VERSION : 0.7
   VAR_INPUT
      FB_Mode : Int;   // Function Block Mode - 0 = HOA Directly Wired to SMC / 1 = HOA Remotely Wired
      MANM : Bool;   // Used only for FB_Mode = 1 / Manual Mode Signal
      AUTM : Bool;   // Used only for FB_Mode = 1 / Auto Mode Signal
      IL : Bool;   // Interlock
      HON : Bool;   // Hand ON
      HOFF : Bool;   // Hand OFF
      SpareIN_1 : Bool;   // Spare
      SRM : Bool;   // Status - Remote Mode Feedback
      SON : Bool;   // Status - On
      SDO : Bool;   // Status - Device Ok
      SCDPA : Bool;   // Status - Cooling Down Period Active
      SESE : Bool;   // Status - Emergency Start Executed
      SGW : Bool;   // Fault - General Warning
      SGF : Bool;   // Fault - General Fault
      EOLO : Bool;   // Event - Overload Operation Fault (I>115%Is)
      EOL : Bool;   // Event - Overload Fault
      EUN : Bool;   // Event - Unbalance Fault
      EOLLP : Bool;   // Event - Overload and Loss of Phase
      ESR : Bool;   // Event - Stalled Rotor
      THFBU : Bool;   // Trip - Hardware Fault Basic Unit
      TMF : Bool;   // Trip - Module Fault
      TEOC : Bool;   // Trip - Execution On-Command
      MC : Int;   // Maximum Current (% of Is)
      IL1 : Int;   // Current of Leg 1 (% of Is)
      IL2 : Int;   // Current of Leg 2 (% of Is)
      IL3 : Int;   // Current of Leg 3 (% of Is)
      RCDP : Int;   // Remaining Cool Down Period
      MOHH : Int;   // Motor Operating Hours High Word
      MOHL : Int;   // Motor Operating Hours Low Word
      LTC : Int;   // Last Trip Current (% of Is)
      "NOT" : Int;   // Number of Overload Trips
      FLA : Real;   // Full Load Amps
   END_VAR
   VAR_OUTPUT
      SpareOUT_1 : Bool;
      Stop_CMD : Bool;   // Stop Command for the Semicode
      Start_CMD : Bool;   // Start Command for the Semicode
      TST : Bool;   // Simocode Test
      EST : Bool;   // Emergency Start
      ERC : Bool;   // Auto Mode / Enable Remote Commands
      RST : Bool;   // Simocode Reset
      SpareOUT_2 : Bool;
      SpareOUT_3 : Bool;
      SpareOUT_4 : Bool;
      SpareOUT_5 : Bool;
      SpareOUT_6 : Bool;
      SpareOUT_7 : Bool;
      SpareOUT_8 : Bool;
      SpareOUT_9 : Bool;
      SpareOUT_10 : Bool;
      SpareOUTW_1 : Int;
      SpareOUTW_2 : Int;
   END_VAR
   VAR
      HMI : Struct
         Controls : Struct
            Start : Bool;
            Stop : Bool;
            Reset : Bool;
            PLCMOHR : Bool;   // PLC Motor Operating Hours Reset
         END_STRUCT;
         Status : Struct
            Mode : Int;   // Simocode Mode
            MotorOperatingHours : Real;   // True Semicode Motor Operating Hours
            DeviceOperatingHours : Real;
            LMOH : Real;   // Last Motor Operating Hours
            RemainingCoolDownPeriod : Int;   // Remaining Cooldown Period
            MaxNumberOLtrips : Int;   // Maximum Number of Overload Trips
            ControlStatusWord : Word;   // Control/Status Information Bits
            MaxCurrent : Real;   // Maximum Current (Is %)
            Current1 : Real;   // Leg 1 Current (Is %)
            Current2 : Real;   // Leg 2 Current (Is %)
            Current3 : Real;   // Leg 3 Current (Is %)
            LastTripCurrent : Real;   // Last Trip Current (% of Is)
            CommandSimocode : Bool;   // Commanding Simocode to Start
         END_STRUCT;
         Config : Struct
            "RemainingCoolDownPeriod.SP" : Int := 300;
            Start_PT : Time := T#500MS;
            Stop_PT : Time := T#500MS;
         END_STRUCT;
         Math : Struct
            MOH1 : DInt;
            MOH2 : Real;
            PLCMOH : Real;   // PLC Motor Operating Hours
            LMOH : Real;
         END_STRUCT;
      END_STRUCT;
      OS : Struct
         RON : Bool;   // Remote / HMI On
         ROFF : Bool;   // Remote / HMI Off
         HON : Bool;   // Hand/Local On
         HOFF : Bool;   // Hand/Local Off
         PLCMOHR : Bool;
         LMOH1 : Bool;
         LMOH2 : Bool;
         RST : Bool;   // Reset Semicode
      END_STRUCT;
      START_CMD_TOF : TOF_TIME;   // Start Semicode
      STOP_CMD_TOF : TOF_TIME;
   END_VAR
   VAR_TEMP
      RMOHH : DInt;
      RMOHL : DInt;
      IL1_Math1 : DInt;
      IL1_Math2 : Real;
      IL1_Math3 : Real;
      IL2_Math1 : DInt;
      IL2_Math2 : Real;
      IL2_Math3 : Real;
      IL3_Math1 : DInt;
      IL3_Math2 : Real;
      IL3_Math3 : Real;
      MC_Math1 : DInt;
      MC_Math2 : Real;
      MC_Math3 : Real;
      LTC_Math1 : DInt;
      LTC_Math2 : Real;
      LTC_Math3 : Real;
      TMOHH : DInt;
      TMOHL : DInt;
      TMOHS : DInt;
   END_VAR
   VAR_TEMP   // added for the SCL form of the ladder/FBD networks
      _w1 : Bool;
      _w2 : Bool;
   END_VAR
BEGIN

REGION Network 1: FB Mode = 0
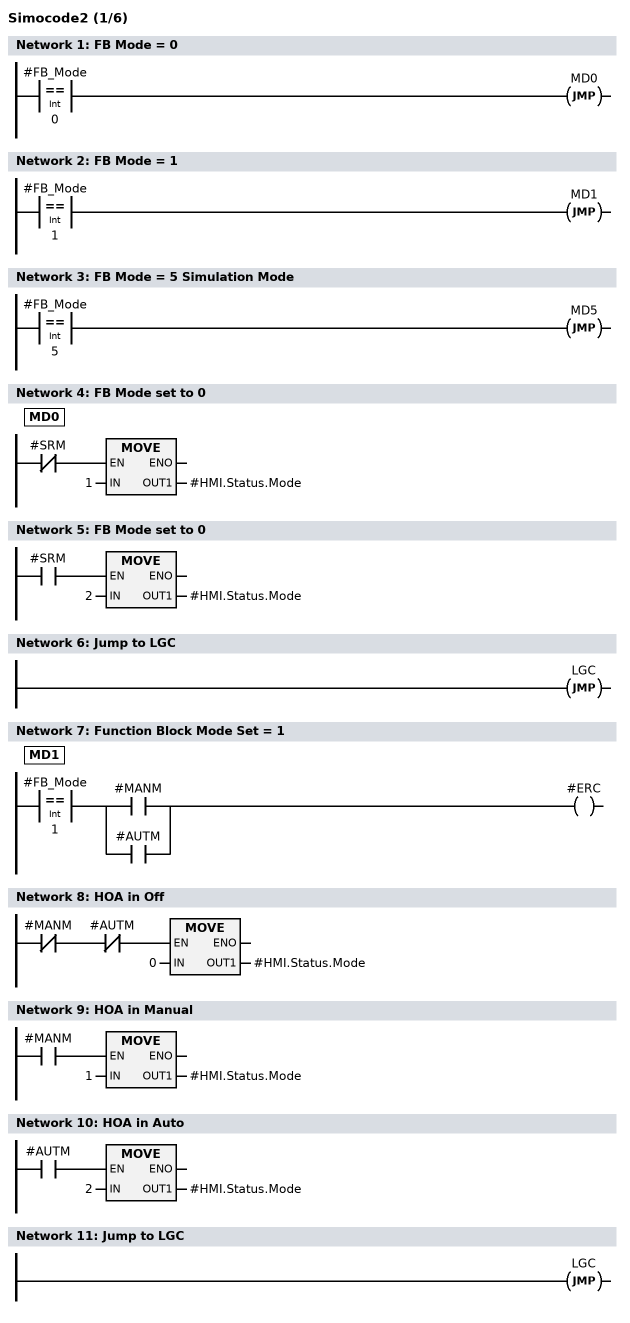
   RUNG wire#powerrail
      { S7_Templates := "SrcType := Int" } EQ_Contact(in1 := #FB_Mode, in2 := 0)
      JumpCoil( MD0 )
   END_RUNG
   // the same network as SCL:
   IF #FB_Mode = 0 THEN GOTO MD0; END_IF;
END_REGION

REGION Network 2: FB Mode = 1
   RUNG wire#powerrail
      { S7_Templates := "SrcType := Int" } EQ_Contact(in1 := #FB_Mode, in2 := 1)
      JumpCoil( MD1 )
   END_RUNG
   // the same network as SCL:
   IF #FB_Mode = 1 THEN GOTO MD1; END_IF;
END_REGION

REGION Network 3: FB Mode = 5 Simulation Mode
   RUNG wire#powerrail
      { S7_Templates := "SrcType := Int" } EQ_Contact(in1 := #FB_Mode, in2 := 5)
      JumpCoil( MD5 )
   END_RUNG
   // the same network as SCL:
   IF #FB_Mode = 5 THEN GOTO MD5; END_IF;
END_REGION

REGION Network 4: FB Mode set to 0
   Label( MD0 )
   RUNG wire#powerrail
      I_Contact( #SRM )
      { S7_GenerateENO := "TRUE" } Move(in := 1, out1 => #HMI.Status.Mode)
   END_RUNG
   // the same network as SCL:
   MD0:
   IF NOT #SRM THEN #HMI.Status.Mode := 1; END_IF;
END_REGION

REGION Network 5: FB Mode set to 0
   RUNG wire#powerrail
      Contact( #SRM )
      { S7_GenerateENO := "TRUE" } Move(in := 2, out1 => #HMI.Status.Mode)
   END_RUNG
   // the same network as SCL:
   IF #SRM THEN #HMI.Status.Mode := 2; END_IF;
END_REGION

REGION Network 6: Jump to LGC
   RUNG wire#powerrail
      JumpCoil( LGC )
   END_RUNG
   // the same network as SCL:
   GOTO LGC;
END_REGION

REGION Network 7: Function Block Mode Set = 1
   Label( MD1 )
   RUNG wire#powerrail
      { S7_Templates := "SrcType := Int" } EQ_Contact(in1 := #FB_Mode, in2 := 1)
      wire#w1
      Contact( #MANM )
      wire#w2
      Coil( #ERC )
   END_RUNG
   RUNG wire#w1
      Contact( #AUTM )
   END_RUNG wire#w2
   // the same network as SCL:
   MD1:
   #ERC := (#FB_Mode = 1) AND (#MANM OR #AUTM);
END_REGION

REGION Network 8: HOA in Off
   RUNG wire#powerrail
      I_Contact( #MANM )
      I_Contact( #AUTM )
      { S7_GenerateENO := "TRUE" } Move(in := 0, out1 => #HMI.Status.Mode)
   END_RUNG
   // the same network as SCL:
   IF NOT #MANM AND NOT #AUTM THEN #HMI.Status.Mode := 0; END_IF;
END_REGION

REGION Network 9: HOA in Manual
   RUNG wire#powerrail
      Contact( #MANM )
      { S7_GenerateENO := "TRUE" } Move(in := 1, out1 => #HMI.Status.Mode)
   END_RUNG
   // the same network as SCL:
   IF #MANM THEN #HMI.Status.Mode := 1; END_IF;
END_REGION

REGION Network 10: HOA in Auto
   RUNG wire#powerrail
      Contact( #AUTM )
      { S7_GenerateENO := "TRUE" } Move(in := 2, out1 => #HMI.Status.Mode)
   END_RUNG
   // the same network as SCL:
   IF #AUTM THEN #HMI.Status.Mode := 2; END_IF;
END_REGION

REGION Network 11: Jump to LGC
   RUNG wire#powerrail
      JumpCoil( LGC )
   END_RUNG
   // the same network as SCL:
   GOTO LGC;
END_REGION

REGION Network 12: FB Mode set to 5
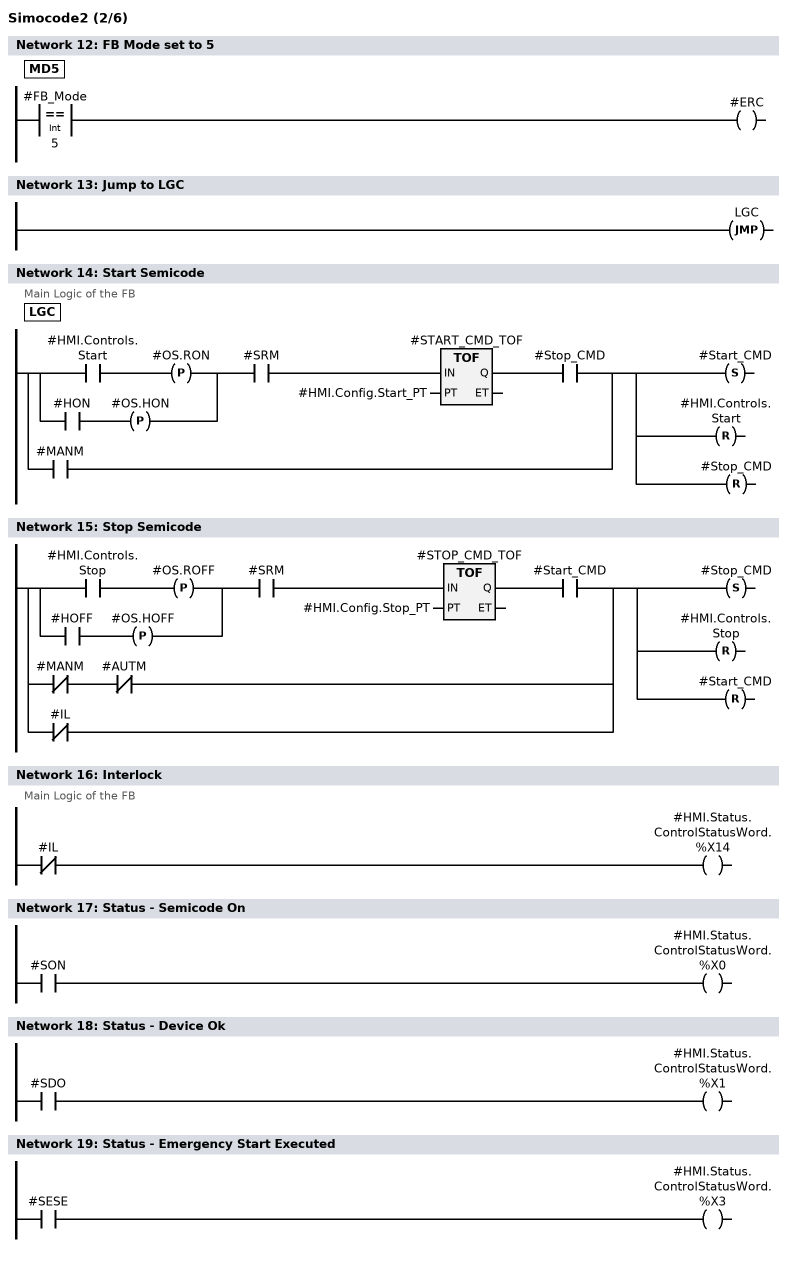
   Label( MD5 )
   RUNG wire#powerrail
      { S7_Templates := "SrcType := Int" } EQ_Contact(in1 := #FB_Mode, in2 := 5)
      Coil( #ERC )
   END_RUNG
   // the same network as SCL:
   MD5:
   #ERC := #FB_Mode = 5;
END_REGION

REGION Network 13: Jump to LGC
   RUNG wire#powerrail
      JumpCoil( LGC )
   END_RUNG
   // the same network as SCL:
   GOTO LGC;
END_REGION

REGION Network 14: Start Semicode
   // Main Logic of the FB
   LGC:
   #_w1 := #HMI.Controls.Start AND NOT #OS.RON;   // rising edge
   #OS.RON := #HMI.Controls.Start;
   #_w2 := #HON AND NOT #OS.HON;   // rising edge
   #OS.HON := #HON;
   #START_CMD_TOF(IN := (#_w1 OR #_w2) AND #SRM, PT := #HMI.Config.Start_PT);   // TOF
   IF (#START_CMD_TOF.Q AND #Stop_CMD) OR #MANM THEN
       #Start_CMD := TRUE;
       #HMI.Controls.Start := FALSE;
       #Stop_CMD := FALSE;
   END_IF;
END_REGION

REGION Network 15: Stop Semicode
   #_w1 := #HMI.Controls.Stop AND NOT #OS.ROFF;   // rising edge
   #OS.ROFF := #HMI.Controls.Stop;
   #_w2 := #HOFF AND NOT #OS.HOFF;   // rising edge
   #OS.HOFF := #HOFF;
   #STOP_CMD_TOF(IN := (#_w1 OR #_w2) AND #SRM, PT := #HMI.Config.Stop_PT);   // TOF
   IF (#STOP_CMD_TOF.Q AND #Start_CMD) OR (NOT #MANM AND NOT #AUTM) OR NOT #IL THEN
       #Stop_CMD := TRUE;
       #HMI.Controls.Stop := FALSE;
       #Start_CMD := FALSE;
   END_IF;
END_REGION

REGION Network 16: Interlock
   // Main Logic of the FB
   RUNG wire#powerrail
      I_Contact( #IL )
      Coil( #HMI.Status.ControlStatusWord.%X14 )
   END_RUNG
   // the same network as SCL:
   #HMI.Status.ControlStatusWord.%X14 := NOT #IL;
END_REGION

REGION Network 17: Status - Semicode On
   RUNG wire#powerrail
      Contact( #SON )
      Coil( #HMI.Status.ControlStatusWord.%X0 )
   END_RUNG
   // the same network as SCL:
   #HMI.Status.ControlStatusWord.%X0 := #SON;
END_REGION

REGION Network 18: Status - Device Ok
   RUNG wire#powerrail
      Contact( #SDO )
      Coil( #HMI.Status.ControlStatusWord.%X1 )
   END_RUNG
   // the same network as SCL:
   #HMI.Status.ControlStatusWord.%X1 := #SDO;
END_REGION

REGION Network 19: Status - Emergency Start Executed
   RUNG wire#powerrail
      Contact( #SESE )
      Coil( #HMI.Status.ControlStatusWord.%X3 )
   END_RUNG
   // the same network as SCL:
   #HMI.Status.ControlStatusWord.%X3 := #SESE;
END_REGION

REGION Network 20: Fault - General Warning
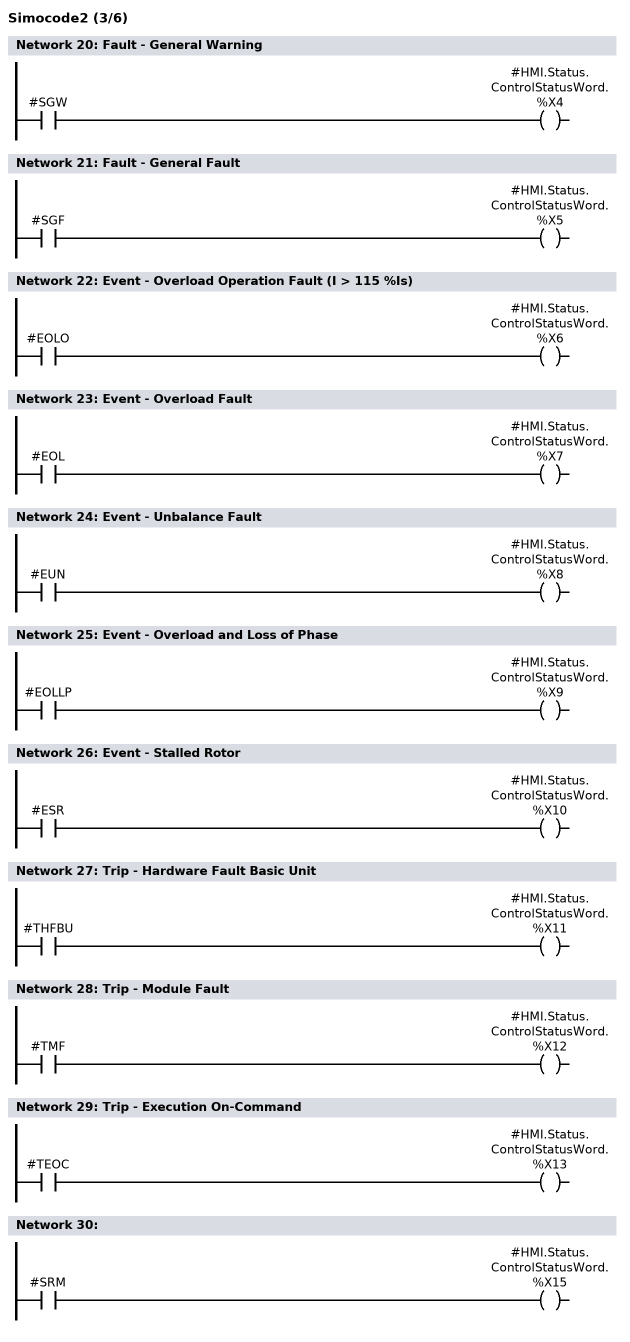
   RUNG wire#powerrail
      Contact( #SGW )
      Coil( #HMI.Status.ControlStatusWord.%X4 )
   END_RUNG
   // the same network as SCL:
   #HMI.Status.ControlStatusWord.%X4 := #SGW;
END_REGION

REGION Network 21: Fault - General Fault
   RUNG wire#powerrail
      Contact( #SGF )
      Coil( #HMI.Status.ControlStatusWord.%X5 )
   END_RUNG
   // the same network as SCL:
   #HMI.Status.ControlStatusWord.%X5 := #SGF;
END_REGION

REGION Network 22: Event - Overload Operation Fault (I > 115 %Is)
   RUNG wire#powerrail
      Contact( #EOLO )
      Coil( #HMI.Status.ControlStatusWord.%X6 )
   END_RUNG
   // the same network as SCL:
   #HMI.Status.ControlStatusWord.%X6 := #EOLO;
END_REGION

REGION Network 23: Event - Overload Fault
   RUNG wire#powerrail
      Contact( #EOL )
      Coil( #HMI.Status.ControlStatusWord.%X7 )
   END_RUNG
   // the same network as SCL:
   #HMI.Status.ControlStatusWord.%X7 := #EOL;
END_REGION

REGION Network 24: Event - Unbalance Fault
   RUNG wire#powerrail
      Contact( #EUN )
      Coil( #HMI.Status.ControlStatusWord.%X8 )
   END_RUNG
   // the same network as SCL:
   #HMI.Status.ControlStatusWord.%X8 := #EUN;
END_REGION

REGION Network 25: Event - Overload and Loss of Phase
   RUNG wire#powerrail
      Contact( #EOLLP )
      Coil( #HMI.Status.ControlStatusWord.%X9 )
   END_RUNG
   // the same network as SCL:
   #HMI.Status.ControlStatusWord.%X9 := #EOLLP;
END_REGION

REGION Network 26: Event - Stalled Rotor
   RUNG wire#powerrail
      Contact( #ESR )
      Coil( #HMI.Status.ControlStatusWord.%X10 )
   END_RUNG
   // the same network as SCL:
   #HMI.Status.ControlStatusWord.%X10 := #ESR;
END_REGION

REGION Network 27: Trip - Hardware Fault Basic Unit
   RUNG wire#powerrail
      Contact( #THFBU )
      Coil( #HMI.Status.ControlStatusWord.%X11 )
   END_RUNG
   // the same network as SCL:
   #HMI.Status.ControlStatusWord.%X11 := #THFBU;
END_REGION

REGION Network 28: Trip - Module Fault
   RUNG wire#powerrail
      Contact( #TMF )
      Coil( #HMI.Status.ControlStatusWord.%X12 )
   END_RUNG
   // the same network as SCL:
   #HMI.Status.ControlStatusWord.%X12 := #TMF;
END_REGION

REGION Network 29: Trip - Execution On-Command
   RUNG wire#powerrail
      Contact( #TEOC )
      Coil( #HMI.Status.ControlStatusWord.%X13 )
   END_RUNG
   // the same network as SCL:
   #HMI.Status.ControlStatusWord.%X13 := #TEOC;
END_REGION

REGION Network 30
   RUNG wire#powerrail
      Contact( #SRM )
      Coil( #HMI.Status.ControlStatusWord.%X15 )
   END_RUNG
   // the same network as SCL:
   #HMI.Status.ControlStatusWord.%X15 := #SRM;
END_REGION

REGION Network 31: Motor Operating Hours
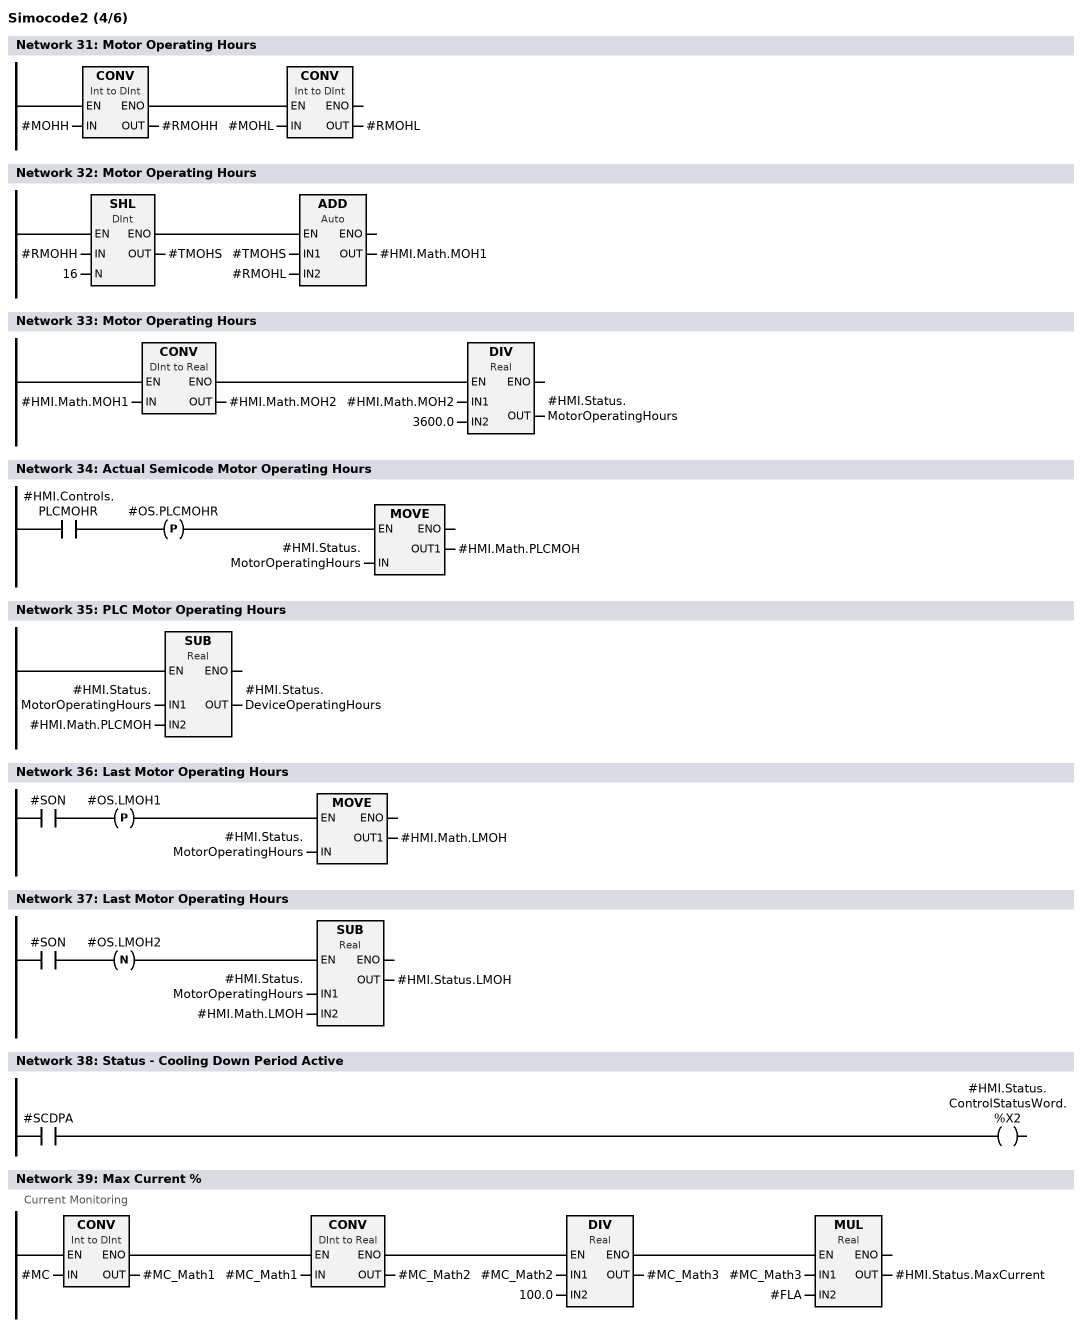
   RUNG wire#powerrail
      { S7_Templates := "[SrcType := Int, DestType := DInt]"; S7_GenerateENO := "TRUE" } Convert(in := #MOHH, out => #RMOHH)
      { S7_Templates := "[SrcType := Int, DestType := DInt]"; S7_GenerateENO := "TRUE" } Convert(in := #MOHL, out => #RMOHL)
   END_RUNG
   // the same network as SCL:
   // ENO of a box is taken as its EN; it also drops when the box reports an error
   #RMOHH := INT_TO_DINT(#MOHH);
   #RMOHL := INT_TO_DINT(#MOHL);
END_REGION

REGION Network 32: Motor Operating Hours
   RUNG wire#powerrail
      { S7_Templates := "SrcType := DInt" } Shl(in := #RMOHH, n := 16, out => #TMOHS)
      Add(in1 := #TMOHS, in2 := #RMOHL, out => #HMI.Math.MOH1)
   END_RUNG
   // the same network as SCL:
   #TMOHS := SHL(IN := #RMOHH, N := 16);
   #HMI.Math.MOH1 := #TMOHS + #RMOHL;
END_REGION

REGION Network 33: Motor Operating Hours
   RUNG wire#powerrail
      { S7_Templates := "[SrcType := DInt, DestType := Real]"; S7_GenerateENO := "TRUE" } Convert(in := #HMI.Math.MOH1, out => #HMI.Math.MOH2)
      { S7_Templates := "SrcType := Real"; S7_GenerateENO := "TRUE" } Div(in1 := #HMI.Math.MOH2, in2 := 3600.0, out => #HMI.Status.MotorOperatingHours)
   END_RUNG
   // the same network as SCL:
   // ENO of a box is taken as its EN; it also drops when the box reports an error
   #HMI.Math.MOH2 := DINT_TO_REAL(#HMI.Math.MOH1);
   #HMI.Status.MotorOperatingHours := #HMI.Math.MOH2 / 3600.0;
END_REGION

REGION Network 34: Actual Semicode Motor Operating Hours
   RUNG wire#powerrail
      Contact( #HMI.Controls.PLCMOHR )
      P_Trig( #OS.PLCMOHR )
      { S7_GenerateENO := "TRUE" } Move(in := #HMI.Status.MotorOperatingHours, out1 => #HMI.Math.PLCMOH)
   END_RUNG
   // the same network as SCL:
   #_w1 := #HMI.Controls.PLCMOHR AND NOT #OS.PLCMOHR;   // rising edge
   #OS.PLCMOHR := #HMI.Controls.PLCMOHR;
   IF #_w1 THEN #HMI.Math.PLCMOH := #HMI.Status.MotorOperatingHours; END_IF;
END_REGION

REGION Network 35: PLC Motor Operating Hours
   RUNG wire#powerrail
      { S7_Templates := "SrcType := Real"; S7_GenerateENO := "TRUE" } Sub(in1 := #HMI.Status.MotorOperatingHours, in2 := #HMI.Math.PLCMOH, out => #HMI.Status.DeviceOperatingHours)
   END_RUNG
   // the same network as SCL:
   #HMI.Status.DeviceOperatingHours := #HMI.Status.MotorOperatingHours - #HMI.Math.PLCMOH;
END_REGION

REGION Network 36: Last Motor Operating Hours
   RUNG wire#powerrail
      Contact( #SON )
      P_Trig( #OS.LMOH1 )
      { S7_GenerateENO := "TRUE" } Move(in := #HMI.Status.MotorOperatingHours, out1 => #HMI.Math.LMOH)
   END_RUNG
   // the same network as SCL:
   #_w1 := #SON AND NOT #OS.LMOH1;   // rising edge
   #OS.LMOH1 := #SON;
   IF #_w1 THEN #HMI.Math.LMOH := #HMI.Status.MotorOperatingHours; END_IF;
END_REGION

REGION Network 37: Last Motor Operating Hours
   RUNG wire#powerrail
      Contact( #SON )
      N_Trig( #OS.LMOH2 )
      { S7_Templates := "SrcType := Real"; S7_GenerateENO := "TRUE" } Sub(in1 := #HMI.Status.MotorOperatingHours, in2 := #HMI.Math.LMOH, out => #HMI.Status.LMOH)
   END_RUNG
   // the same network as SCL:
   #_w1 := NOT #SON AND #OS.LMOH2;   // falling edge
   #OS.LMOH2 := #SON;
   IF #_w1 THEN #HMI.Status.LMOH := #HMI.Status.MotorOperatingHours - #HMI.Math.LMOH; END_IF;
END_REGION

REGION Network 38: Status - Cooling Down Period Active
   RUNG wire#powerrail
      Contact( #SCDPA )
      Coil( #HMI.Status.ControlStatusWord.%X2 )
   END_RUNG
   // the same network as SCL:
   #HMI.Status.ControlStatusWord.%X2 := #SCDPA;
END_REGION

REGION Network 39: Max Current %
   // Current Monitoring
   RUNG wire#powerrail
      { S7_Templates := "[SrcType := Int, DestType := DInt]"; S7_GenerateENO := "TRUE" } Convert(in := #MC, out => #MC_Math1)
      { S7_Templates := "[SrcType := DInt, DestType := Real]"; S7_GenerateENO := "TRUE" } Convert(in := #MC_Math1, out => #MC_Math2)
      { S7_Templates := "SrcType := Real"; S7_GenerateENO := "TRUE" } Div(in1 := #MC_Math2, in2 := 100.0, out => #MC_Math3)
      { S7_Templates := "SrcType := Real"; S7_GenerateENO := "TRUE" } Mul(in1 := #MC_Math3, in2 := #FLA, out => #HMI.Status.MaxCurrent)
   END_RUNG
   // the same network as SCL:
   // ENO of a box is taken as its EN; it also drops when the box reports an error
   #MC_Math1 := INT_TO_DINT(#MC);
   #MC_Math2 := DINT_TO_REAL(#MC_Math1);
   #MC_Math3 := #MC_Math2 / 100.0;
   #HMI.Status.MaxCurrent := #MC_Math3 * #FLA;
END_REGION

REGION Network 40: L1 Current %
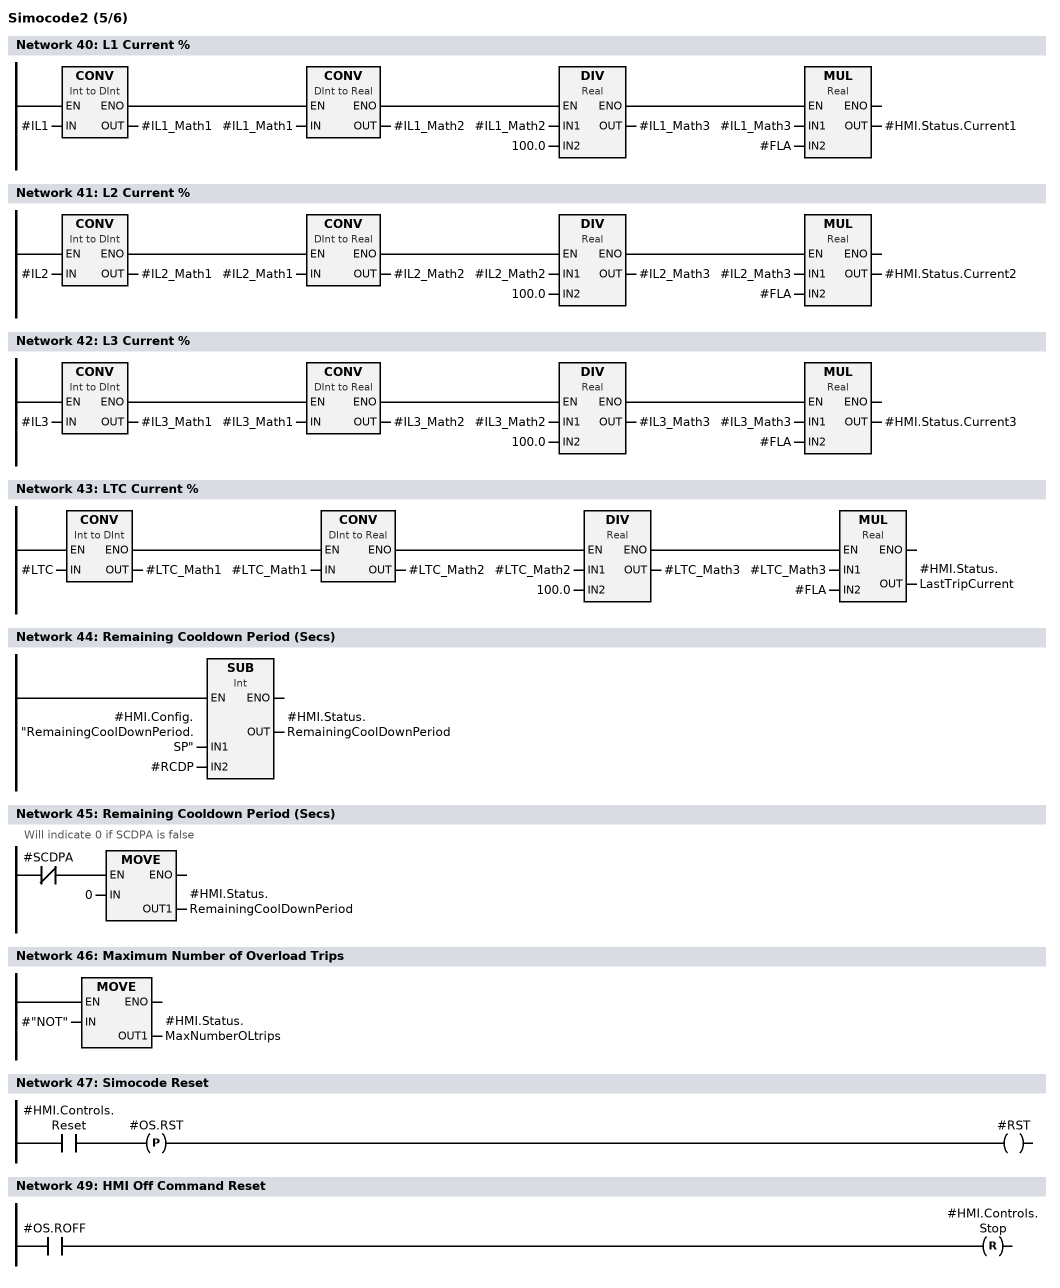
   RUNG wire#powerrail
      { S7_Templates := "[SrcType := Int, DestType := DInt]"; S7_GenerateENO := "TRUE" } Convert(in := #IL1, out => #IL1_Math1)
      { S7_Templates := "[SrcType := DInt, DestType := Real]"; S7_GenerateENO := "TRUE" } Convert(in := #IL1_Math1, out => #IL1_Math2)
      { S7_Templates := "SrcType := Real"; S7_GenerateENO := "TRUE" } Div(in1 := #IL1_Math2, in2 := 100.0, out => #IL1_Math3)
      { S7_Templates := "SrcType := Real"; S7_GenerateENO := "TRUE" } Mul(in1 := #IL1_Math3, in2 := #FLA, out => #HMI.Status.Current1)
   END_RUNG
   // the same network as SCL:
   // ENO of a box is taken as its EN; it also drops when the box reports an error
   #IL1_Math1 := INT_TO_DINT(#IL1);
   #IL1_Math2 := DINT_TO_REAL(#IL1_Math1);
   #IL1_Math3 := #IL1_Math2 / 100.0;
   #HMI.Status.Current1 := #IL1_Math3 * #FLA;
END_REGION

REGION Network 41: L2 Current %
   RUNG wire#powerrail
      { S7_Templates := "[SrcType := Int, DestType := DInt]"; S7_GenerateENO := "TRUE" } Convert(in := #IL2, out => #IL2_Math1)
      { S7_Templates := "[SrcType := DInt, DestType := Real]"; S7_GenerateENO := "TRUE" } Convert(in := #IL2_Math1, out => #IL2_Math2)
      { S7_Templates := "SrcType := Real"; S7_GenerateENO := "TRUE" } Div(in1 := #IL2_Math2, in2 := 100.0, out => #IL2_Math3)
      { S7_Templates := "SrcType := Real"; S7_GenerateENO := "TRUE" } Mul(in1 := #IL2_Math3, in2 := #FLA, out => #HMI.Status.Current2)
   END_RUNG
   // the same network as SCL:
   // ENO of a box is taken as its EN; it also drops when the box reports an error
   #IL2_Math1 := INT_TO_DINT(#IL2);
   #IL2_Math2 := DINT_TO_REAL(#IL2_Math1);
   #IL2_Math3 := #IL2_Math2 / 100.0;
   #HMI.Status.Current2 := #IL2_Math3 * #FLA;
END_REGION

REGION Network 42: L3 Current %
   RUNG wire#powerrail
      { S7_Templates := "[SrcType := Int, DestType := DInt]"; S7_GenerateENO := "TRUE" } Convert(in := #IL3, out => #IL3_Math1)
      { S7_Templates := "[SrcType := DInt, DestType := Real]"; S7_GenerateENO := "TRUE" } Convert(in := #IL3_Math1, out => #IL3_Math2)
      { S7_Templates := "SrcType := Real"; S7_GenerateENO := "TRUE" } Div(in1 := #IL3_Math2, in2 := 100.0, out => #IL3_Math3)
      { S7_Templates := "SrcType := Real"; S7_GenerateENO := "TRUE" } Mul(in1 := #IL3_Math3, in2 := #FLA, out => #HMI.Status.Current3)
   END_RUNG
   // the same network as SCL:
   // ENO of a box is taken as its EN; it also drops when the box reports an error
   #IL3_Math1 := INT_TO_DINT(#IL3);
   #IL3_Math2 := DINT_TO_REAL(#IL3_Math1);
   #IL3_Math3 := #IL3_Math2 / 100.0;
   #HMI.Status.Current3 := #IL3_Math3 * #FLA;
END_REGION

REGION Network 43: LTC Current %
   RUNG wire#powerrail
      { S7_Templates := "[SrcType := Int, DestType := DInt]"; S7_GenerateENO := "TRUE" } Convert(in := #LTC, out => #LTC_Math1)
      { S7_Templates := "[SrcType := DInt, DestType := Real]"; S7_GenerateENO := "TRUE" } Convert(in := #LTC_Math1, out => #LTC_Math2)
      { S7_Templates := "SrcType := Real"; S7_GenerateENO := "TRUE" } Div(in1 := #LTC_Math2, in2 := 100.0, out => #LTC_Math3)
      { S7_Templates := "SrcType := Real"; S7_GenerateENO := "TRUE" } Mul(in1 := #LTC_Math3, in2 := #FLA, out => #HMI.Status.LastTripCurrent)
   END_RUNG
   // the same network as SCL:
   // ENO of a box is taken as its EN; it also drops when the box reports an error
   #LTC_Math1 := INT_TO_DINT(#LTC);
   #LTC_Math2 := DINT_TO_REAL(#LTC_Math1);
   #LTC_Math3 := #LTC_Math2 / 100.0;
   #HMI.Status.LastTripCurrent := #LTC_Math3 * #FLA;
END_REGION

REGION Network 44: Remaining Cooldown Period (Secs)
   RUNG wire#powerrail
      { S7_Templates := "SrcType := Int"; S7_GenerateENO := "TRUE" } Sub(in1 := #HMI.Config."RemainingCoolDownPeriod.SP", in2 := #RCDP, out => #HMI.Status.RemainingCoolDownPeriod)
   END_RUNG
   // the same network as SCL:
   #HMI.Status.RemainingCoolDownPeriod := #HMI.Config."RemainingCoolDownPeriod.SP" - #RCDP;
END_REGION

REGION Network 45: Remaining Cooldown Period (Secs)
   // Will indicate 0 if SCDPA is false
   RUNG wire#powerrail
      I_Contact( #SCDPA )
      { S7_GenerateENO := "TRUE" } Move(in := 0, out1 => #HMI.Status.RemainingCoolDownPeriod)
   END_RUNG
   // the same network as SCL:
   IF NOT #SCDPA THEN #HMI.Status.RemainingCoolDownPeriod := 0; END_IF;
END_REGION

REGION Network 46: Maximum Number of Overload Trips
   RUNG wire#powerrail
      { S7_GenerateENO := "TRUE" } Move(in := #"NOT", out1 => #HMI.Status.MaxNumberOLtrips)
   END_RUNG
   // the same network as SCL:
   #HMI.Status.MaxNumberOLtrips := #"NOT";
END_REGION

REGION Network 47: Simocode Reset
   RUNG wire#powerrail
      Contact( #HMI.Controls.Reset )
      P_Trig( #OS.RST )
      Coil( #RST )
   END_RUNG
   // the same network as SCL:
   #_w1 := #HMI.Controls.Reset AND NOT #OS.RST;   // rising edge
   #OS.RST := #HMI.Controls.Reset;
   #RST := #_w1;
END_REGION

REGION Network 48: HMI On Command Reset
   // HMI Command Resets
END_REGION

REGION Network 49: HMI Off Command Reset
   RUNG wire#powerrail
      Contact( #OS.ROFF )
      R_Coil( #HMI.Controls.Stop )
   END_RUNG
   // the same network as SCL:
   IF #OS.ROFF THEN #HMI.Controls.Stop := FALSE; END_IF;
END_REGION

REGION Network 50: Simocode Reset PB Clear
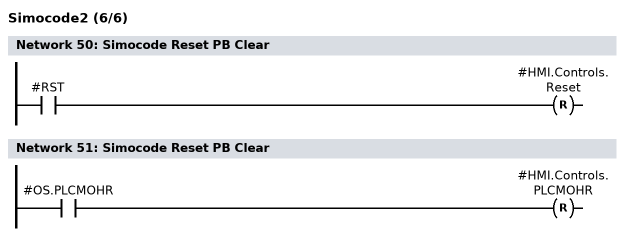
   RUNG wire#powerrail
      Contact( #RST )
      R_Coil( #HMI.Controls.Reset )
   END_RUNG
   // the same network as SCL:
   IF #RST THEN #HMI.Controls.Reset := FALSE; END_IF;
END_REGION

REGION Network 51: Simocode Reset PB Clear
   RUNG wire#powerrail
      Contact( #OS.PLCMOHR )
      R_Coil( #HMI.Controls.PLCMOHR )
   END_RUNG
   // the same network as SCL:
   IF #OS.PLCMOHR THEN #HMI.Controls.PLCMOHR := FALSE; END_IF;
END_REGION
END_FUNCTION_BLOCK

// folder: 1}Library/Split Range

FUNCTION_BLOCK "Split Range 'V'"   // FB7, LAD
{ S7_Optimized_Access := 'TRUE' }
VERSION : 0.1
   VAR_INPUT
      "PID Output" : Real;   // Output of the controller
      RangeX : Real;   // range desired from 0 to X
      RangeY : Real;   // range desired from X to Y
   END_VAR
   VAR_OUTPUT
      "Range1.Q" : Int;
      "Range2.Q" : Int;
   END_VAR
   VAR_TEMP
      div1 : Real;
      out1 : Real;
      rawout1 : Real;
      "scaling.a3" : Real;
      deadband : Real;
      range2pdb : Real;
      newmvi : Real;
      newmviabs : Real;
      div2 : Real;
      out2 : Real;
      rawout2 : Real;
      dintRound : DInt;
      intOutput : Int;
      test1 : Real;
   END_VAR
   VAR_TEMP   // added for the SCL form of the ladder/FBD networks
      _w1 : Bool;
   END_VAR
BEGIN

REGION Network 1: Split range X
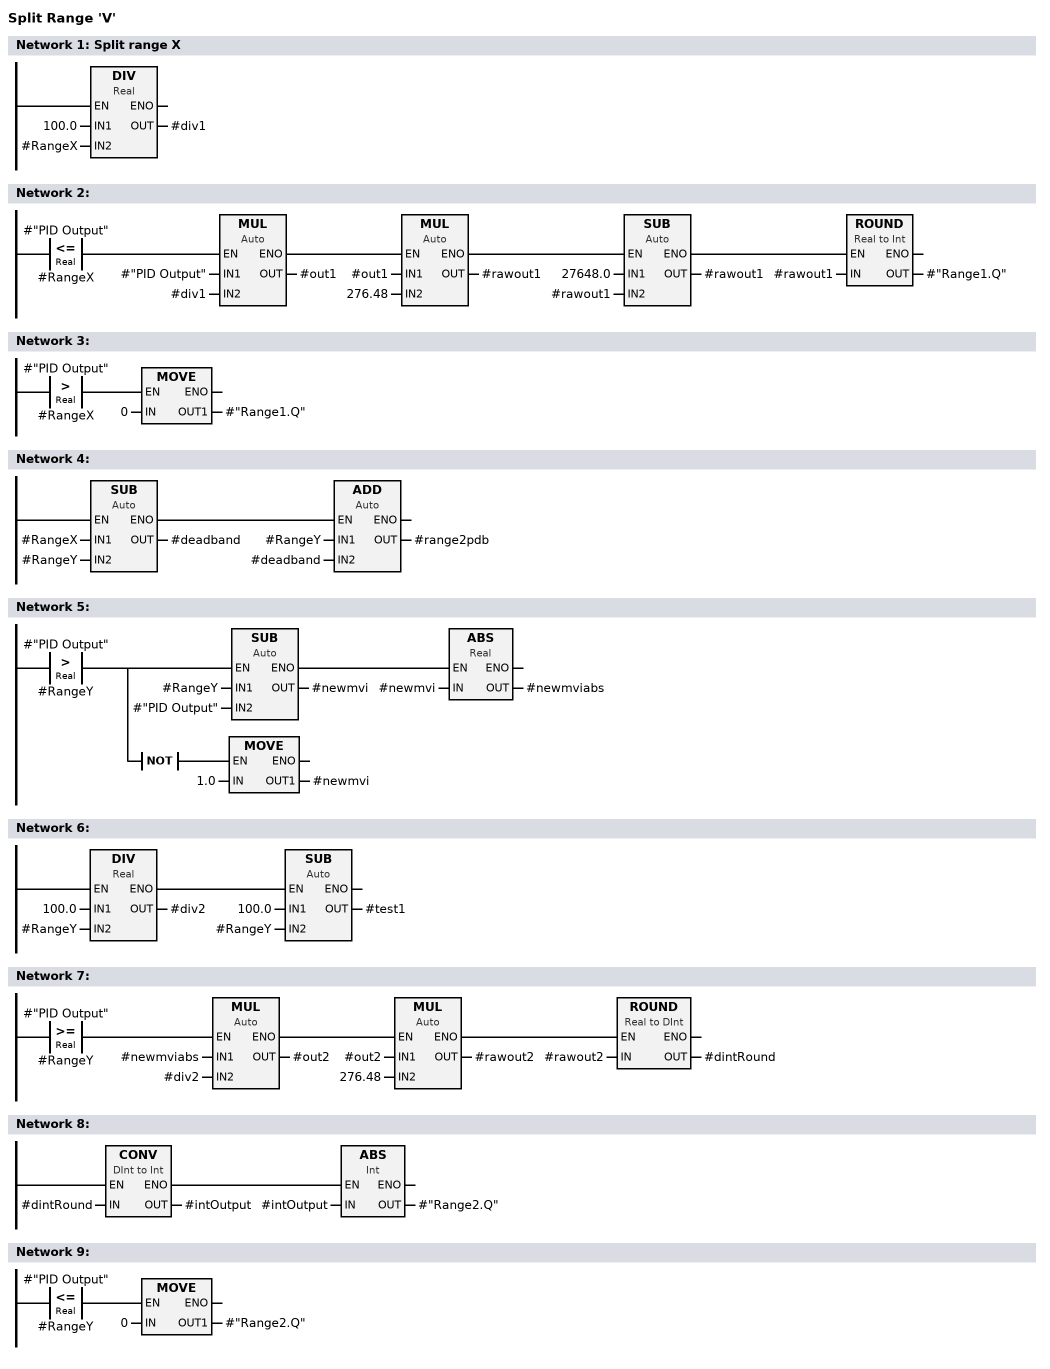
   RUNG wire#powerrail
      { S7_Templates := "SrcType := Real" } Div(in1 := 100.0, in2 := #RangeX, out => #div1)
   END_RUNG
   // the same network as SCL:
   #div1 := 100.0 / #RangeX;
END_REGION

REGION Network 2
   RUNG wire#powerrail
      { S7_Templates := "SrcType := Real" } LE_Contact(in1 := #"PID Output", in2 := #RangeX)
      Mul(in1 := #"PID Output", in2 := #div1, out => #out1)
      Mul(in1 := #out1, in2 := 276.48, out => #rawout1)
      Sub(in1 := 27648.0, in2 := #rawout1, out => #rawout1)
      { S7_Templates := "[SrcType := Real, DestType := Int]" } Round(in := #rawout1, out => #"Range1.Q")
   END_RUNG
   // the same network as SCL:
   IF #"PID Output" <= #RangeX THEN
       #out1 := #"PID Output" * #div1;
       #rawout1 := #out1 * 276.48;
       #rawout1 := 27648.0 - #rawout1;
       #"Range1.Q" := ROUND(#rawout1);
   END_IF;
END_REGION

REGION Network 3
   RUNG wire#powerrail
      { S7_Templates := "SrcType := Real" } GT_Contact(in1 := #"PID Output", in2 := #RangeX)
      Move(in := 0, out1 => #"Range1.Q")
   END_RUNG
   // the same network as SCL:
   IF #"PID Output" > #RangeX THEN #"Range1.Q" := 0; END_IF;
END_REGION

REGION Network 4
   RUNG wire#powerrail
      Sub(in1 := #RangeX, in2 := #RangeY, out => #deadband)
      Add(in1 := #RangeY, in2 := #deadband, out => #range2pdb)
   END_RUNG
   // the same network as SCL:
   #deadband := #RangeX - #RangeY;
   #range2pdb := #RangeY + #deadband;
END_REGION

REGION Network 5
   RUNG wire#powerrail
      { S7_Templates := "SrcType := Real" } GT_Contact(in1 := #"PID Output", in2 := #RangeY)
      wire#w1
      Sub(in1 := #RangeY, in2 := #"PID Output", out => #newmvi)
      { S7_Templates := "SrcType := Real" } Abs(in := #newmvi, out => #newmviabs)
   END_RUNG
   RUNG wire#w1
      Not()
      Move(in := 1.0, out1 => #newmvi)
   END_RUNG
   // the same network as SCL:
   #_w1 := #"PID Output" > #RangeY;
   IF #_w1 THEN
       #newmvi := #RangeY - #"PID Output";
       #newmviabs := ABS(#newmvi);
   END_IF;
   IF NOT #_w1 THEN #newmvi := 1.0; END_IF;
END_REGION

REGION Network 6
   RUNG wire#powerrail
      { S7_Templates := "SrcType := Real" } Div(in1 := 100.0, in2 := #RangeY, out => #div2)
      Sub(in1 := 100.0, in2 := #RangeY, out => #test1)
   END_RUNG
   // the same network as SCL:
   #div2 := 100.0 / #RangeY;
   #test1 := 100.0 - #RangeY;
END_REGION

REGION Network 7
   RUNG wire#powerrail
      { S7_Templates := "SrcType := Real" } GE_Contact(in1 := #"PID Output", in2 := #RangeY)
      Mul(in1 := #newmviabs, in2 := #div2, out => #out2)
      Mul(in1 := #out2, in2 := 276.48, out => #rawout2)
      { S7_Templates := "[SrcType := Real, DestType := DInt]" } Round(in := #rawout2, out => #dintRound)
   END_RUNG
   // the same network as SCL:
   IF #"PID Output" >= #RangeY THEN
       #out2 := #newmviabs * #div2;
       #rawout2 := #out2 * 276.48;
       #dintRound := ROUND(#rawout2);
   END_IF;
END_REGION

REGION Network 8
   RUNG wire#powerrail
      { S7_Templates := "[SrcType := DInt, DestType := Int]" } Convert(in := #dintRound, out => #intOutput)
      { S7_Templates := "SrcType := Int" } Abs(in := #intOutput, out => #"Range2.Q")
   END_RUNG
   // the same network as SCL:
   #intOutput := DINT_TO_INT(#dintRound);
   #"Range2.Q" := ABS(#intOutput);
END_REGION
